REGION Network 21
   RUNG wire#powerrail
      Contact( "Carrier_21_Status.9" )
      Coil( "EMS".Carrier[21].SDC_IN.EncoderCommFault )
   END_RUNG
   // the same network as SCL:
   "EMS".Carrier[21].SDC_IN.EncoderCommFault := "Carrier_21_Status.9";
END_REGION

REGION Network 22
   RUNG wire#powerrail
      Contact( "Carrier_21_Status.10" )
      Coil( "EMS".Carrier[21].SDC_IN.DriveCommFault )
   END_RUNG
   // the same network as SCL:
   "EMS".Carrier[21].SDC_IN.DriveCommFault := "Carrier_21_Status.10";
END_REGION

REGION Network 23
   RUNG wire#powerrail
      Contact( "Carrier_21_Status.11" )
      Coil( "EMS".Carrier[21].SDC_IN.HMICommFault )
   END_RUNG
   // the same network as SCL:
   "EMS".Carrier[21].SDC_IN.HMICommFault := "Carrier_21_Status.11";
END_REGION

REGION Network 24
   RUNG wire#powerrail
      Contact( "Carrier_21_Status.2" )
      Coil( "EMS".Carrier[21].SDC_IN.AutoMode )
   END_RUNG
   RUNG wire#powerrail
      Contact( "Carrier_21_Status.1" )
      Coil( "EMS".Carrier[21].SDC_IN.ManualMode )
   END_RUNG
   // the same network as SCL:
   "EMS".Carrier[21].SDC_IN.AutoMode := "Carrier_21_Status.2";
   "EMS".Carrier[21].SDC_IN.ManualMode := "Carrier_21_Status.1";
END_REGION

REGION Network 25
   Label( C21_Comm_Fault )
   RUNG wire#powerrail
      Coil( "SectionComment" )
   END_RUNG
   // the same network as SCL:
   C21_Comm_Fault:
   "SectionComment" := TRUE;
END_REGION

REGION Network 26
   // **********************************************************************************************************************
   // 
   // Carrier 22 I-Device Data Transfer Interlocks from Carrier to SDC
   // 
   // **********************************************************************************************************************
   RUNG wire#powerrail
      Coil( "SectionComment" )
   END_RUNG
   // the same network as SCL:
   "SectionComment" := TRUE;
END_REGION

REGION Network 27
   RUNG wire#powerrail
      { S7_Templates := "SrcType := Word" } NE_Contact(in1 := "Carrier_22_CarrierNumber", in2 := 0)
      Move(in := "Carrier_22_CarrierNumber", out1 => "EMS".Carrier[22].SDC_IN.CarrierNumber)
   END_RUNG
   // the same network as SCL:
   IF "Carrier_22_CarrierNumber" <> 0 THEN
       "EMS".Carrier[22].SDC_IN.CarrierNumber := "Carrier_22_CarrierNumber";
   END_IF;
END_REGION

REGION Network 28
   RUNG wire#powerrail
      { S7_Templates := "SrcType := DWord" } NE_Contact(in1 := "Carrier_22_CarrierPosition", in2 := 0)
      Move(in := "Carrier_22_CarrierPosition", out1 => "EMS".Carrier[22].SDC_IN.CarrierPosition)
   END_RUNG
   // the same network as SCL:
   IF "Carrier_22_CarrierPosition" <> 0 THEN
       "EMS".Carrier[22].SDC_IN.CarrierPosition := "Carrier_22_CarrierPosition";
   END_IF;
END_REGION

REGION Network 29
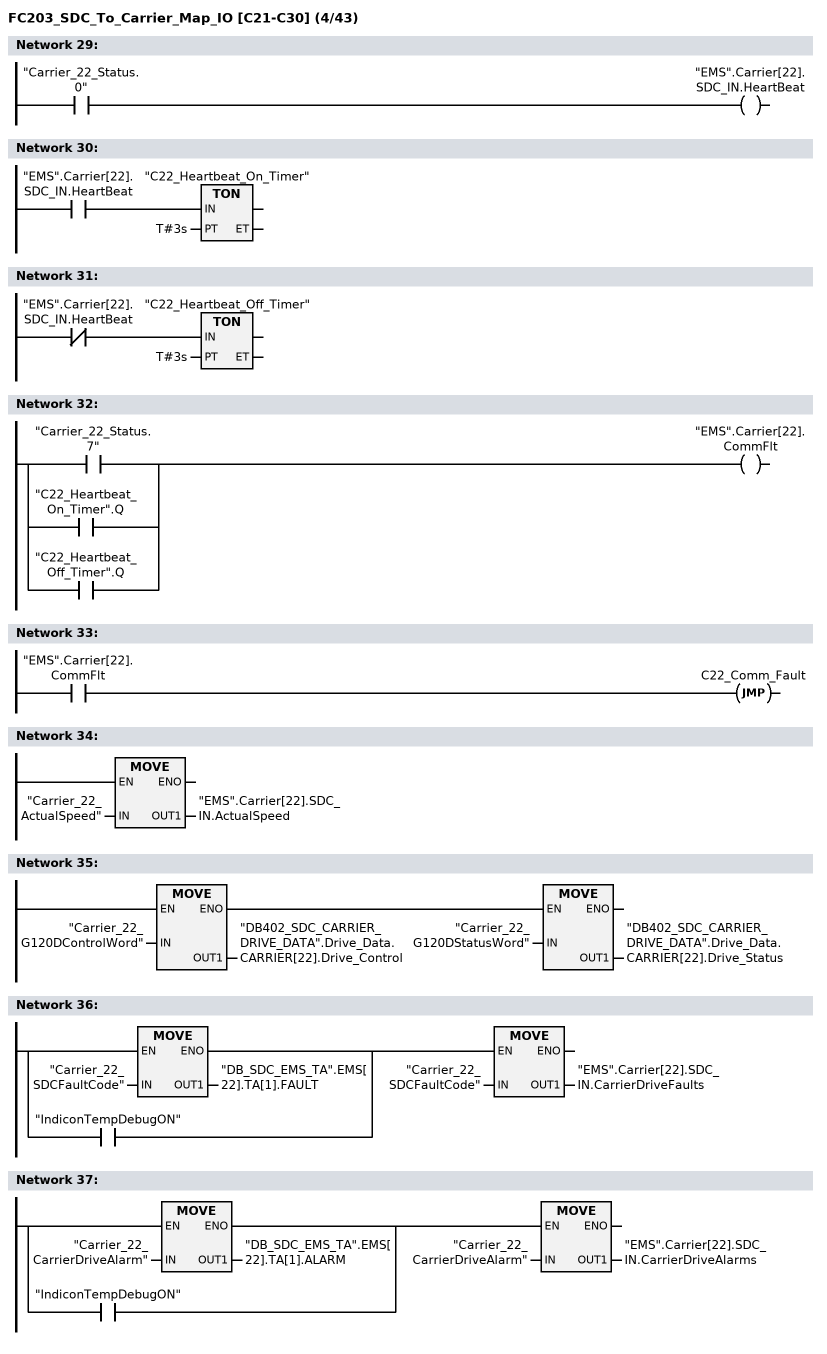
   RUNG wire#powerrail
      Contact( "Carrier_22_Status.0" )
      Coil( "EMS".Carrier[22].SDC_IN.HeartBeat )
   END_RUNG
   // the same network as SCL:
   "EMS".Carrier[22].SDC_IN.HeartBeat := "Carrier_22_Status.0";
END_REGION

REGION Network 30
   "C22_Heartbeat_On_Timer".TON(IN := "EMS".Carrier[22].SDC_IN.HeartBeat, PT := T#3s);
END_REGION

REGION Network 31
   "C22_Heartbeat_Off_Timer".TON(IN := NOT "EMS".Carrier[22].SDC_IN.HeartBeat, PT := T#3s);
END_REGION

REGION Network 32
   RUNG wire#powerrail
      Contact( "Carrier_22_Status.7" )
      wire#w1
      Coil( "EMS".Carrier[22].CommFlt )
   END_RUNG
   RUNG wire#powerrail
      Contact( "C22_Heartbeat_On_Timer".Q )
   END_RUNG wire#w1
   RUNG wire#powerrail
      Contact( "C22_Heartbeat_Off_Timer".Q )
   END_RUNG wire#w1
   // the same network as SCL:
   "EMS".Carrier[22].CommFlt := "Carrier_22_Status.7" OR "C22_Heartbeat_On_Timer".Q OR "C22_Heartbeat_Off_Timer".Q;
END_REGION

REGION Network 33
   RUNG wire#powerrail
      Contact( "EMS".Carrier[22].CommFlt )
      JumpCoil( C22_Comm_Fault )
   END_RUNG
   // the same network as SCL:
   IF "EMS".Carrier[22].CommFlt THEN GOTO C22_Comm_Fault; END_IF;
END_REGION

REGION Network 34
   RUNG wire#powerrail
      Move(in := "Carrier_22_ActualSpeed", out1 => "EMS".Carrier[22].SDC_IN.ActualSpeed)
   END_RUNG
   // the same network as SCL:
   "EMS".Carrier[22].SDC_IN.ActualSpeed := "Carrier_22_ActualSpeed";
END_REGION

REGION Network 35
   RUNG wire#powerrail
      Move(in := "Carrier_22_G120DControlWord", out1 => "DB402_SDC_CARRIER_DRIVE_DATA".Drive_Data.CARRIER[22].Drive_Control)
      Move(in := "Carrier_22_G120DStatusWord", out1 => "DB402_SDC_CARRIER_DRIVE_DATA".Drive_Data.CARRIER[22].Drive_Status)
   END_RUNG
   // the same network as SCL:
   "DB402_SDC_CARRIER_DRIVE_DATA".Drive_Data.CARRIER[22].Drive_Control := "Carrier_22_G120DControlWord";
   "DB402_SDC_CARRIER_DRIVE_DATA".Drive_Data.CARRIER[22].Drive_Status := "Carrier_22_G120DStatusWord";
END_REGION

REGION Network 36
   RUNG wire#powerrail
      Move(in := "Carrier_22_SDCFaultCode", out1 => "DB_SDC_EMS_TA".EMS[22].TA[1].FAULT)
      wire#w1
      Move(in := "Carrier_22_SDCFaultCode", out1 => "EMS".Carrier[22].SDC_IN.CarrierDriveFaults)
   END_RUNG
   RUNG wire#powerrail
      Contact( "IndiconTempDebugON" )
   END_RUNG wire#w1
   // the same network as SCL:
   "DB_SDC_EMS_TA".EMS[22].TA[1].FAULT := "Carrier_22_SDCFaultCode";
   IF TRUE OR "IndiconTempDebugON" THEN
       "EMS".Carrier[22].SDC_IN.CarrierDriveFaults := "Carrier_22_SDCFaultCode";
   END_IF;
END_REGION

REGION Network 37
   RUNG wire#powerrail
      Move(in := "Carrier_22_CarrierDriveAlarm", out1 => "DB_SDC_EMS_TA".EMS[22].TA[1].ALARM)
      wire#w1
      Move(in := "Carrier_22_CarrierDriveAlarm", out1 => "EMS".Carrier[22].SDC_IN.CarrierDriveAlarms)
   END_RUNG
   RUNG wire#powerrail
      Contact( "IndiconTempDebugON" )
   END_RUNG wire#w1
   // the same network as SCL:
   "DB_SDC_EMS_TA".EMS[22].TA[1].ALARM := "Carrier_22_CarrierDriveAlarm";
   IF TRUE OR "IndiconTempDebugON" THEN
       "EMS".Carrier[22].SDC_IN.CarrierDriveAlarms := "Carrier_22_CarrierDriveAlarm";
   END_IF;
END_REGION

REGION Network 38
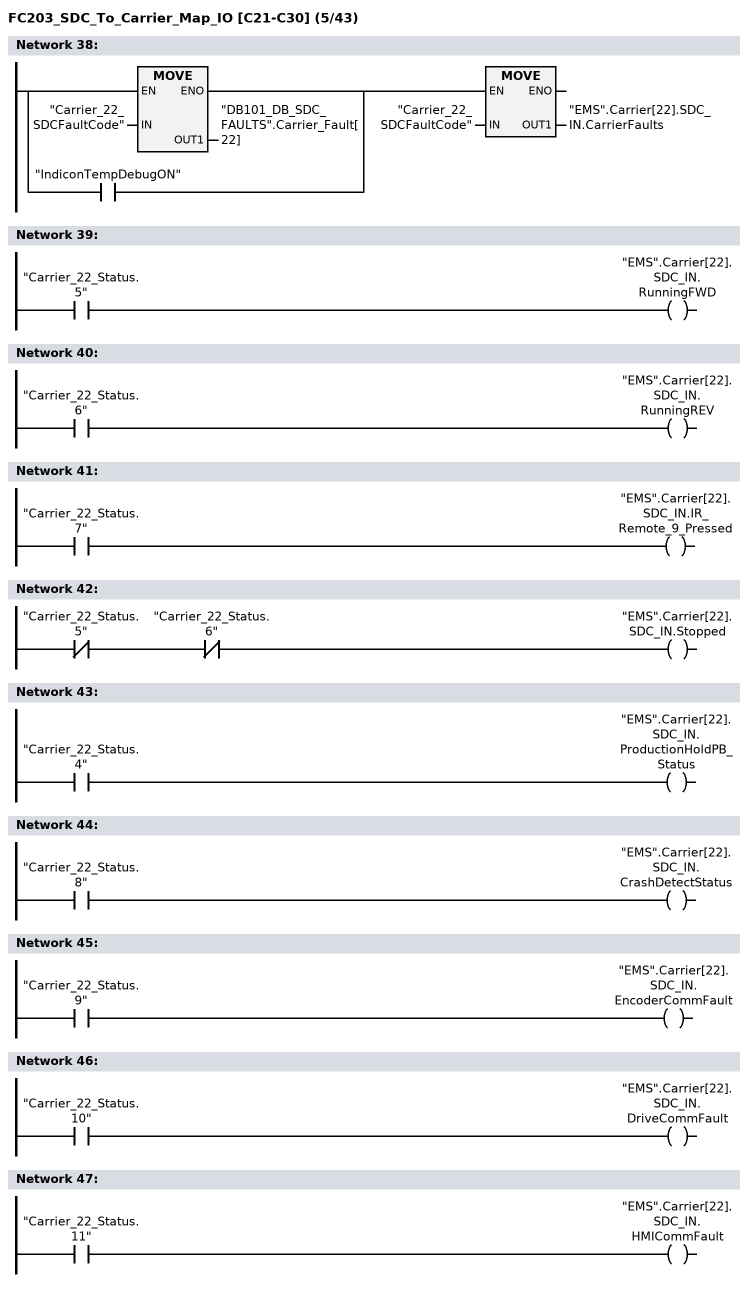
   RUNG wire#powerrail
      Move(in := "Carrier_22_SDCFaultCode", out1 => "DB101_DB_SDC_FAULTS".Carrier_Fault[22])
      wire#w1
      Move(in := "Carrier_22_SDCFaultCode", out1 => "EMS".Carrier[22].SDC_IN.CarrierFaults)
   END_RUNG
   RUNG wire#powerrail
      Contact( "IndiconTempDebugON" )
   END_RUNG wire#w1
   // the same network as SCL:
   "DB101_DB_SDC_FAULTS".Carrier_Fault[22] := "Carrier_22_SDCFaultCode";
   IF TRUE OR "IndiconTempDebugON" THEN
       "EMS".Carrier[22].SDC_IN.CarrierFaults := "Carrier_22_SDCFaultCode";
   END_IF;
END_REGION

REGION Network 39
   RUNG wire#powerrail
      Contact( "Carrier_22_Status.5" )
      Coil( "EMS".Carrier[22].SDC_IN.RunningFWD )
   END_RUNG
   // the same network as SCL:
   "EMS".Carrier[22].SDC_IN.RunningFWD := "Carrier_22_Status.5";
END_REGION

REGION Network 40
   RUNG wire#powerrail
      Contact( "Carrier_22_Status.6" )
      Coil( "EMS".Carrier[22].SDC_IN.RunningREV )
   END_RUNG
   // the same network as SCL:
   "EMS".Carrier[22].SDC_IN.RunningREV := "Carrier_22_Status.6";
END_REGION

REGION Network 41
   RUNG wire#powerrail
      Contact( "Carrier_22_Status.7" )
      Coil( "EMS".Carrier[22].SDC_IN.IR_Remote_9_Pressed )
   END_RUNG
   // the same network as SCL:
   "EMS".Carrier[22].SDC_IN.IR_Remote_9_Pressed := "Carrier_22_Status.7";
END_REGION

REGION Network 42
   RUNG wire#powerrail
      I_Contact( "Carrier_22_Status.5" )
      I_Contact( "Carrier_22_Status.6" )
      Coil( "EMS".Carrier[22].SDC_IN.Stopped )
   END_RUNG
   // the same network as SCL:
   "EMS".Carrier[22].SDC_IN.Stopped := NOT "Carrier_22_Status.5" AND NOT "Carrier_22_Status.6";
END_REGION

REGION Network 43
   RUNG wire#powerrail
      Contact( "Carrier_22_Status.4" )
      Coil( "EMS".Carrier[22].SDC_IN.ProductionHoldPB_Status )
   END_RUNG
   // the same network as SCL:
   "EMS".Carrier[22].SDC_IN.ProductionHoldPB_Status := "Carrier_22_Status.4";
END_REGION

REGION Network 44
   RUNG wire#powerrail
      Contact( "Carrier_22_Status.8" )
      Coil( "EMS".Carrier[22].SDC_IN.CrashDetectStatus )
   END_RUNG
   // the same network as SCL:
   "EMS".Carrier[22].SDC_IN.CrashDetectStatus := "Carrier_22_Status.8";
END_REGION

REGION Network 45
   RUNG wire#powerrail
      Contact( "Carrier_22_Status.9" )
      Coil( "EMS".Carrier[22].SDC_IN.EncoderCommFault )
   END_RUNG
   // the same network as SCL:
   "EMS".Carrier[22].SDC_IN.EncoderCommFault := "Carrier_22_Status.9";
END_REGION

REGION Network 46
   RUNG wire#powerrail
      Contact( "Carrier_22_Status.10" )
      Coil( "EMS".Carrier[22].SDC_IN.DriveCommFault )
   END_RUNG
   // the same network as SCL:
   "EMS".Carrier[22].SDC_IN.DriveCommFault := "Carrier_22_Status.10";
END_REGION

REGION Network 47
   RUNG wire#powerrail
      Contact( "Carrier_22_Status.11" )
      Coil( "EMS".Carrier[22].SDC_IN.HMICommFault )
   END_RUNG
   // the same network as SCL:
   "EMS".Carrier[22].SDC_IN.HMICommFault := "Carrier_22_Status.11";
END_REGION

REGION Network 48
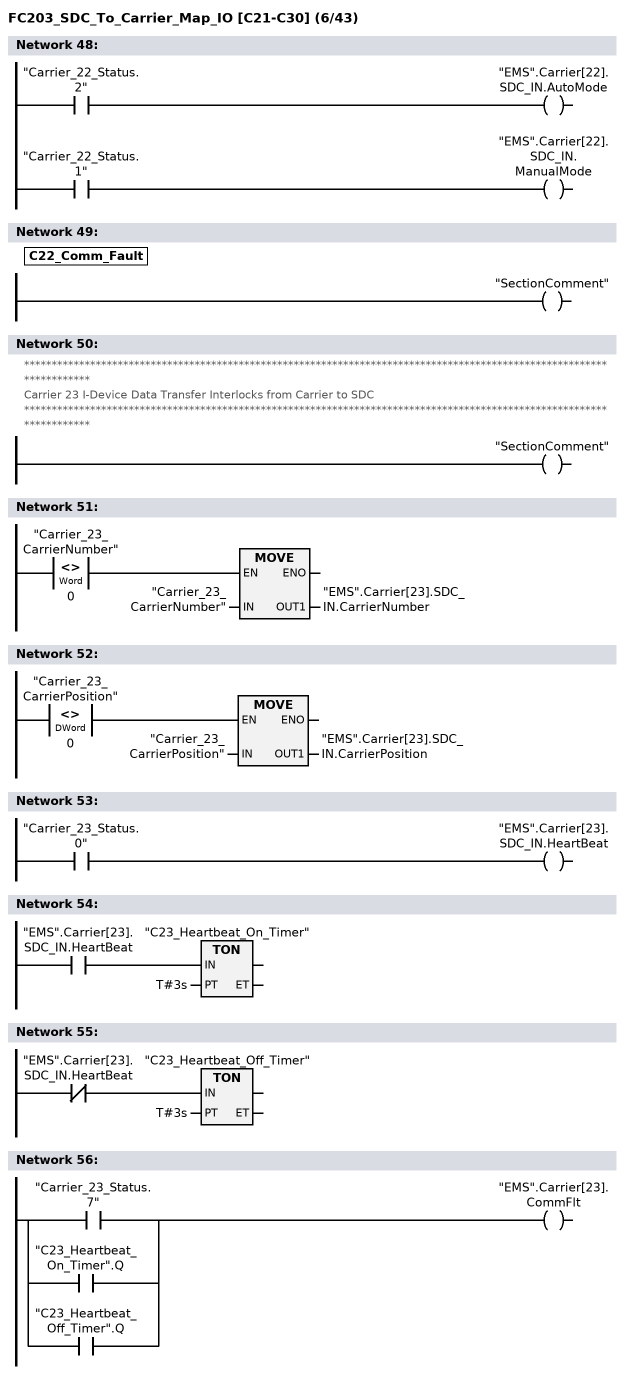
   RUNG wire#powerrail
      Contact( "Carrier_22_Status.2" )
      Coil( "EMS".Carrier[22].SDC_IN.AutoMode )
   END_RUNG
   RUNG wire#powerrail
      Contact( "Carrier_22_Status.1" )
      Coil( "EMS".Carrier[22].SDC_IN.ManualMode )
   END_RUNG
   // the same network as SCL:
   "EMS".Carrier[22].SDC_IN.AutoMode := "Carrier_22_Status.2";
   "EMS".Carrier[22].SDC_IN.ManualMode := "Carrier_22_Status.1";
END_REGION

REGION Network 49
   Label( C22_Comm_Fault )
   RUNG wire#powerrail
      Coil( "SectionComment" )
   END_RUNG
   // the same network as SCL:
   C22_Comm_Fault:
   "SectionComment" := TRUE;
END_REGION

REGION Network 50
   // **********************************************************************************************************************
   // 
   // Carrier 23 I-Device Data Transfer Interlocks from Carrier to SDC
   // 
   // **********************************************************************************************************************
   RUNG wire#powerrail
      Coil( "SectionComment" )
   END_RUNG
   // the same network as SCL:
   "SectionComment" := TRUE;
END_REGION

REGION Network 51
   RUNG wire#powerrail
      { S7_Templates := "SrcType := Word" } NE_Contact(in1 := "Carrier_23_CarrierNumber", in2 := 0)
      Move(in := "Carrier_23_CarrierNumber", out1 => "EMS".Carrier[23].SDC_IN.CarrierNumber)
   END_RUNG
   // the same network as SCL:
   IF "Carrier_23_CarrierNumber" <> 0 THEN
       "EMS".Carrier[23].SDC_IN.CarrierNumber := "Carrier_23_CarrierNumber";
   END_IF;
END_REGION

REGION Network 52
   RUNG wire#powerrail
      { S7_Templates := "SrcType := DWord" } NE_Contact(in1 := "Carrier_23_CarrierPosition", in2 := 0)
      Move(in := "Carrier_23_CarrierPosition", out1 => "EMS".Carrier[23].SDC_IN.CarrierPosition)
   END_RUNG
   // the same network as SCL:
   IF "Carrier_23_CarrierPosition" <> 0 THEN
       "EMS".Carrier[23].SDC_IN.CarrierPosition := "Carrier_23_CarrierPosition";
   END_IF;
END_REGION

REGION Network 53
   RUNG wire#powerrail
      Contact( "Carrier_23_Status.0" )
      Coil( "EMS".Carrier[23].SDC_IN.HeartBeat )
   END_RUNG
   // the same network as SCL:
   "EMS".Carrier[23].SDC_IN.HeartBeat := "Carrier_23_Status.0";
END_REGION

REGION Network 54
   "C23_Heartbeat_On_Timer".TON(IN := "EMS".Carrier[23].SDC_IN.HeartBeat, PT := T#3s);
END_REGION

REGION Network 55
   "C23_Heartbeat_Off_Timer".TON(IN := NOT "EMS".Carrier[23].SDC_IN.HeartBeat, PT := T#3s);
END_REGION

REGION Network 56
   RUNG wire#powerrail
      Contact( "Carrier_23_Status.7" )
      wire#w1
      Coil( "EMS".Carrier[23].CommFlt )
   END_RUNG
   RUNG wire#powerrail
      Contact( "C23_Heartbeat_On_Timer".Q )
   END_RUNG wire#w1
   RUNG wire#powerrail
      Contact( "C23_Heartbeat_Off_Timer".Q )
   END_RUNG wire#w1
   // the same network as SCL:
   "EMS".Carrier[23].CommFlt := "Carrier_23_Status.7" OR "C23_Heartbeat_On_Timer".Q OR "C23_Heartbeat_Off_Timer".Q;
END_REGION

REGION Network 57
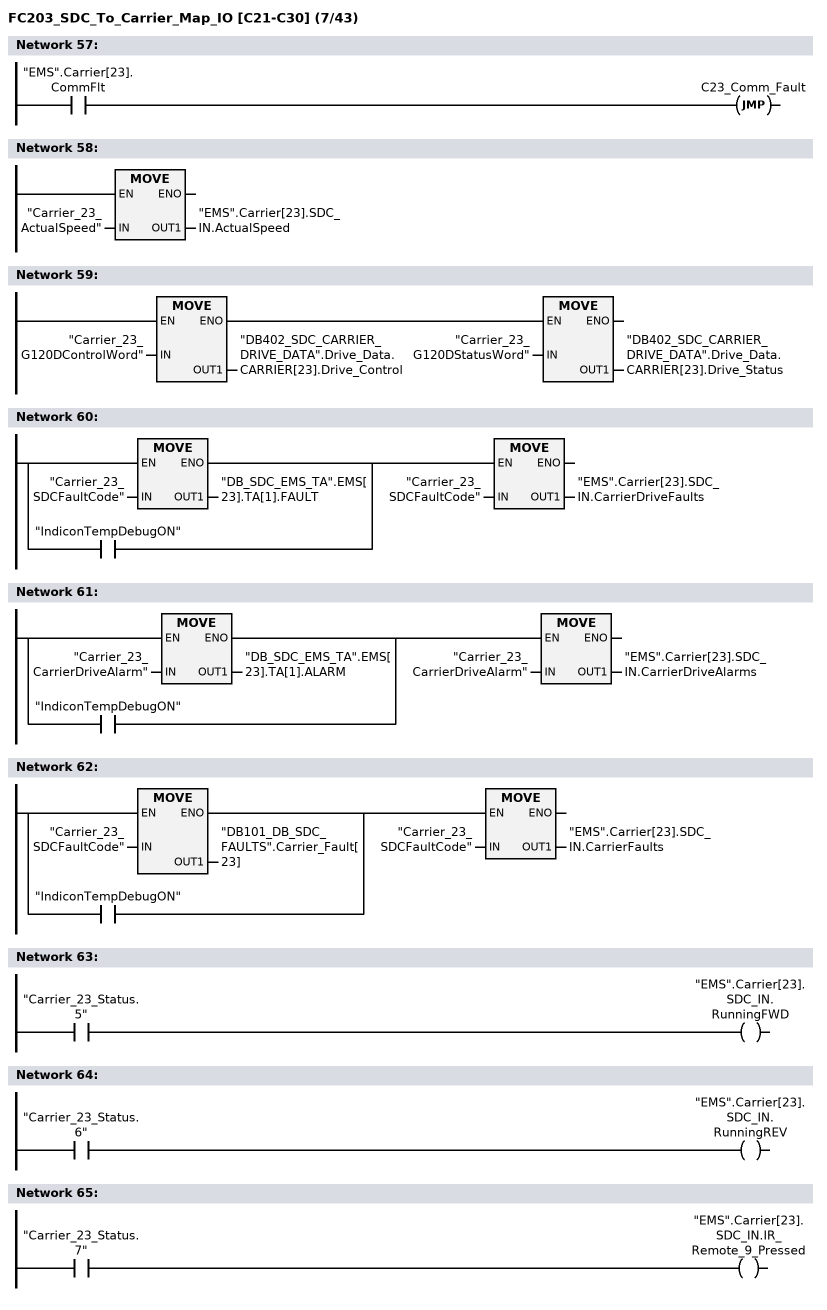
   RUNG wire#powerrail
      Contact( "EMS".Carrier[23].CommFlt )
      JumpCoil( C23_Comm_Fault )
   END_RUNG
   // the same network as SCL:
   IF "EMS".Carrier[23].CommFlt THEN GOTO C23_Comm_Fault; END_IF;
END_REGION

REGION Network 58
   RUNG wire#powerrail
      Move(in := "Carrier_23_ActualSpeed", out1 => "EMS".Carrier[23].SDC_IN.ActualSpeed)
   END_RUNG
   // the same network as SCL:
   "EMS".Carrier[23].SDC_IN.ActualSpeed := "Carrier_23_ActualSpeed";
END_REGION

REGION Network 59
   RUNG wire#powerrail
      Move(in := "Carrier_23_G120DControlWord", out1 => "DB402_SDC_CARRIER_DRIVE_DATA".Drive_Data.CARRIER[23].Drive_Control)
      Move(in := "Carrier_23_G120DStatusWord", out1 => "DB402_SDC_CARRIER_DRIVE_DATA".Drive_Data.CARRIER[23].Drive_Status)
   END_RUNG
   // the same network as SCL:
   "DB402_SDC_CARRIER_DRIVE_DATA".Drive_Data.CARRIER[23].Drive_Control := "Carrier_23_G120DControlWord";
   "DB402_SDC_CARRIER_DRIVE_DATA".Drive_Data.CARRIER[23].Drive_Status := "Carrier_23_G120DStatusWord";
END_REGION

REGION Network 60
   RUNG wire#powerrail
      Move(in := "Carrier_23_SDCFaultCode", out1 => "DB_SDC_EMS_TA".EMS[23].TA[1].FAULT)
      wire#w1
      Move(in := "Carrier_23_SDCFaultCode", out1 => "EMS".Carrier[23].SDC_IN.CarrierDriveFaults)
   END_RUNG
   RUNG wire#powerrail
      Contact( "IndiconTempDebugON" )
   END_RUNG wire#w1
   // the same network as SCL:
   "DB_SDC_EMS_TA".EMS[23].TA[1].FAULT := "Carrier_23_SDCFaultCode";
   IF TRUE OR "IndiconTempDebugON" THEN
       "EMS".Carrier[23].SDC_IN.CarrierDriveFaults := "Carrier_23_SDCFaultCode";
   END_IF;
END_REGION

REGION Network 61
   RUNG wire#powerrail
      Move(in := "Carrier_23_CarrierDriveAlarm", out1 => "DB_SDC_EMS_TA".EMS[23].TA[1].ALARM)
      wire#w1
      Move(in := "Carrier_23_CarrierDriveAlarm", out1 => "EMS".Carrier[23].SDC_IN.CarrierDriveAlarms)
   END_RUNG
   RUNG wire#powerrail
      Contact( "IndiconTempDebugON" )
   END_RUNG wire#w1
   // the same network as SCL:
   "DB_SDC_EMS_TA".EMS[23].TA[1].ALARM := "Carrier_23_CarrierDriveAlarm";
   IF TRUE OR "IndiconTempDebugON" THEN
       "EMS".Carrier[23].SDC_IN.CarrierDriveAlarms := "Carrier_23_CarrierDriveAlarm";
   END_IF;
END_REGION

REGION Network 62
   RUNG wire#powerrail
      Move(in := "Carrier_23_SDCFaultCode", out1 => "DB101_DB_SDC_FAULTS".Carrier_Fault[23])
      wire#w1
      Move(in := "Carrier_23_SDCFaultCode", out1 => "EMS".Carrier[23].SDC_IN.CarrierFaults)
   END_RUNG
   RUNG wire#powerrail
      Contact( "IndiconTempDebugON" )
   END_RUNG wire#w1
   // the same network as SCL:
   "DB101_DB_SDC_FAULTS".Carrier_Fault[23] := "Carrier_23_SDCFaultCode";
   IF TRUE OR "IndiconTempDebugON" THEN
       "EMS".Carrier[23].SDC_IN.CarrierFaults := "Carrier_23_SDCFaultCode";
   END_IF;
END_REGION

REGION Network 63
   RUNG wire#powerrail
      Contact( "Carrier_23_Status.5" )
      Coil( "EMS".Carrier[23].SDC_IN.RunningFWD )
   END_RUNG
   // the same network as SCL:
   "EMS".Carrier[23].SDC_IN.RunningFWD := "Carrier_23_Status.5";
END_REGION

REGION Network 64
   RUNG wire#powerrail
      Contact( "Carrier_23_Status.6" )
      Coil( "EMS".Carrier[23].SDC_IN.RunningREV )
   END_RUNG
   // the same network as SCL:
   "EMS".Carrier[23].SDC_IN.RunningREV := "Carrier_23_Status.6";
END_REGION

REGION Network 65
   RUNG wire#powerrail
      Contact( "Carrier_23_Status.7" )
      Coil( "EMS".Carrier[23].SDC_IN.IR_Remote_9_Pressed )
   END_RUNG
   // the same network as SCL:
   "EMS".Carrier[23].SDC_IN.IR_Remote_9_Pressed := "Carrier_23_Status.7";
END_REGION

REGION Network 66
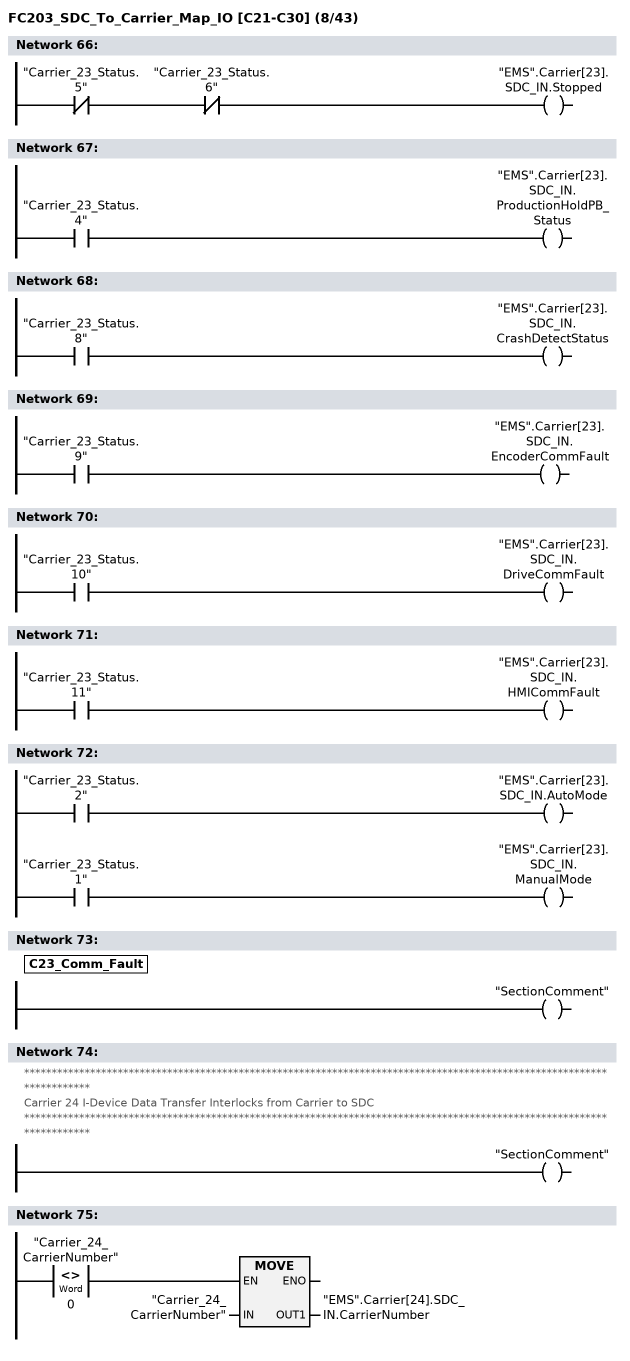
   RUNG wire#powerrail
      I_Contact( "Carrier_23_Status.5" )
      I_Contact( "Carrier_23_Status.6" )
      Coil( "EMS".Carrier[23].SDC_IN.Stopped )
   END_RUNG
   // the same network as SCL:
   "EMS".Carrier[23].SDC_IN.Stopped := NOT "Carrier_23_Status.5" AND NOT "Carrier_23_Status.6";
END_REGION

REGION Network 67
   RUNG wire#powerrail
      Contact( "Carrier_23_Status.4" )
      Coil( "EMS".Carrier[23].SDC_IN.ProductionHoldPB_Status )
   END_RUNG
   // the same network as SCL:
   "EMS".Carrier[23].SDC_IN.ProductionHoldPB_Status := "Carrier_23_Status.4";
END_REGION

REGION Network 68
   RUNG wire#powerrail
      Contact( "Carrier_23_Status.8" )
      Coil( "EMS".Carrier[23].SDC_IN.CrashDetectStatus )
   END_RUNG
   // the same network as SCL:
   "EMS".Carrier[23].SDC_IN.CrashDetectStatus := "Carrier_23_Status.8";
END_REGION

REGION Network 69
   RUNG wire#powerrail
      Contact( "Carrier_23_Status.9" )
      Coil( "EMS".Carrier[23].SDC_IN.EncoderCommFault )
   END_RUNG
   // the same network as SCL:
   "EMS".Carrier[23].SDC_IN.EncoderCommFault := "Carrier_23_Status.9";
END_REGION

REGION Network 70
   RUNG wire#powerrail
      Contact( "Carrier_23_Status.10" )
      Coil( "EMS".Carrier[23].SDC_IN.DriveCommFault )
   END_RUNG
   // the same network as SCL:
   "EMS".Carrier[23].SDC_IN.DriveCommFault := "Carrier_23_Status.10";
END_REGION

REGION Network 71
   RUNG wire#powerrail
      Contact( "Carrier_23_Status.11" )
      Coil( "EMS".Carrier[23].SDC_IN.HMICommFault )
   END_RUNG
   // the same network as SCL:
   "EMS".Carrier[23].SDC_IN.HMICommFault := "Carrier_23_Status.11";
END_REGION

REGION Network 72
   RUNG wire#powerrail
      Contact( "Carrier_23_Status.2" )
      Coil( "EMS".Carrier[23].SDC_IN.AutoMode )
   END_RUNG
   RUNG wire#powerrail
      Contact( "Carrier_23_Status.1" )
      Coil( "EMS".Carrier[23].SDC_IN.ManualMode )
   END_RUNG
   // the same network as SCL:
   "EMS".Carrier[23].SDC_IN.AutoMode := "Carrier_23_Status.2";
   "EMS".Carrier[23].SDC_IN.ManualMode := "Carrier_23_Status.1";
END_REGION

REGION Network 73
   Label( C23_Comm_Fault )
   RUNG wire#powerrail
      Coil( "SectionComment" )
   END_RUNG
   // the same network as SCL:
   C23_Comm_Fault:
   "SectionComment" := TRUE;
END_REGION

REGION Network 74
   // **********************************************************************************************************************
   // 
   // Carrier 24 I-Device Data Transfer Interlocks from Carrier to SDC
   // 
   // **********************************************************************************************************************
   RUNG wire#powerrail
      Coil( "SectionComment" )
   END_RUNG
   // the same network as SCL:
   "SectionComment" := TRUE;
END_REGION

REGION Network 75
   RUNG wire#powerrail
      { S7_Templates := "SrcType := Word" } NE_Contact(in1 := "Carrier_24_CarrierNumber", in2 := 0)
      Move(in := "Carrier_24_CarrierNumber", out1 => "EMS".Carrier[24].SDC_IN.CarrierNumber)
   END_RUNG
   // the same network as SCL:
   IF "Carrier_24_CarrierNumber" <> 0 THEN
       "EMS".Carrier[24].SDC_IN.CarrierNumber := "Carrier_24_CarrierNumber";
   END_IF;
END_REGION

REGION Network 76
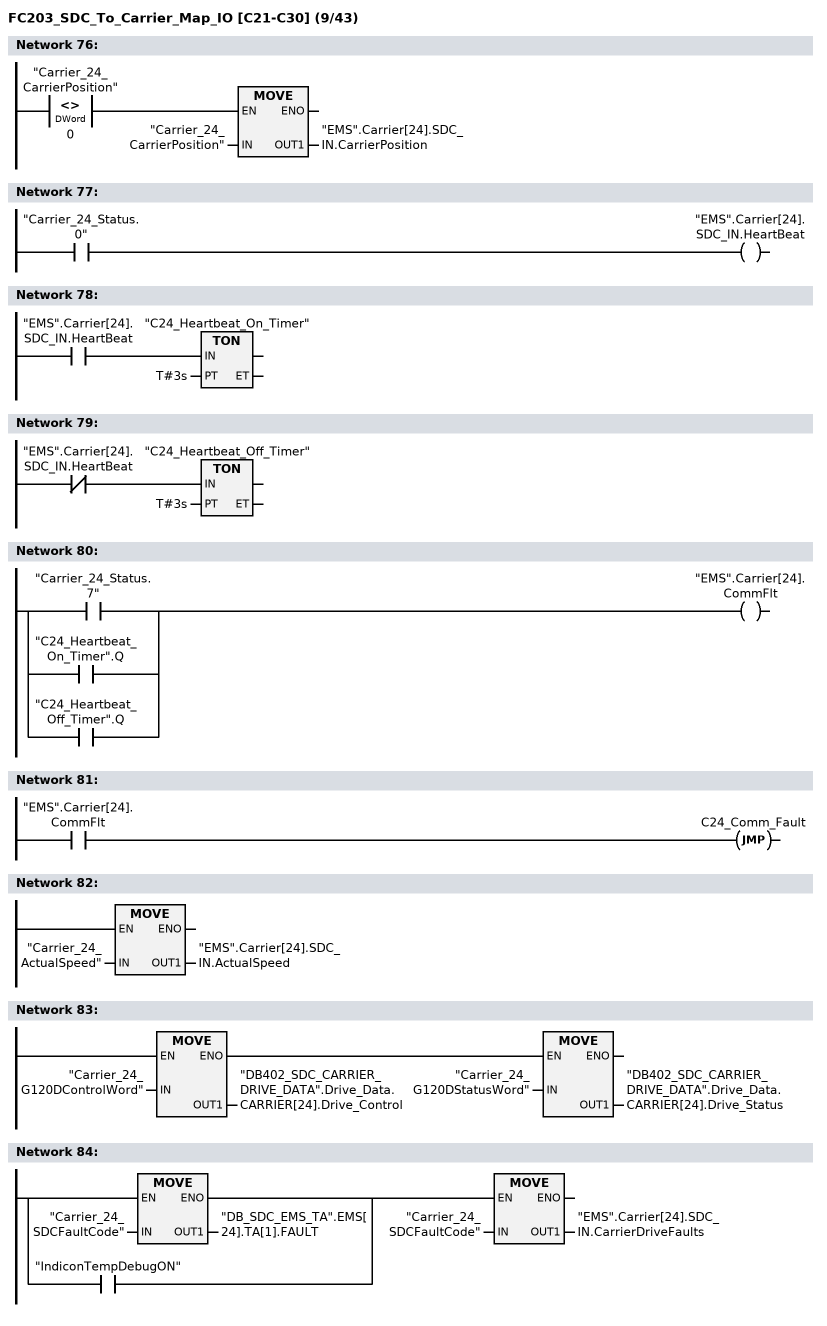
   RUNG wire#powerrail
      { S7_Templates := "SrcType := DWord" } NE_Contact(in1 := "Carrier_24_CarrierPosition", in2 := 0)
      Move(in := "Carrier_24_CarrierPosition", out1 => "EMS".Carrier[24].SDC_IN.CarrierPosition)
   END_RUNG
   // the same network as SCL:
   IF "Carrier_24_CarrierPosition" <> 0 THEN
       "EMS".Carrier[24].SDC_IN.CarrierPosition := "Carrier_24_CarrierPosition";
   END_IF;
END_REGION

REGION Network 77
   RUNG wire#powerrail
      Contact( "Carrier_24_Status.0" )
      Coil( "EMS".Carrier[24].SDC_IN.HeartBeat )
   END_RUNG
   // the same network as SCL:
   "EMS".Carrier[24].SDC_IN.HeartBeat := "Carrier_24_Status.0";
END_REGION

REGION Network 78
   "C24_Heartbeat_On_Timer".TON(IN := "EMS".Carrier[24].SDC_IN.HeartBeat, PT := T#3s);
END_REGION

REGION Network 79
   "C24_Heartbeat_Off_Timer".TON(IN := NOT "EMS".Carrier[24].SDC_IN.HeartBeat, PT := T#3s);
END_REGION

REGION Network 80
   RUNG wire#powerrail
      Contact( "Carrier_24_Status.7" )
      wire#w1
      Coil( "EMS".Carrier[24].CommFlt )
   END_RUNG
   RUNG wire#powerrail
      Contact( "C24_Heartbeat_On_Timer".Q )
   END_RUNG wire#w1
   RUNG wire#powerrail
      Contact( "C24_Heartbeat_Off_Timer".Q )
   END_RUNG wire#w1
   // the same network as SCL:
   "EMS".Carrier[24].CommFlt := "Carrier_24_Status.7" OR "C24_Heartbeat_On_Timer".Q OR "C24_Heartbeat_Off_Timer".Q;
END_REGION

REGION Network 81
   RUNG wire#powerrail
      Contact( "EMS".Carrier[24].CommFlt )
      JumpCoil( C24_Comm_Fault )
   END_RUNG
   // the same network as SCL:
   IF "EMS".Carrier[24].CommFlt THEN GOTO C24_Comm_Fault; END_IF;
END_REGION

REGION Network 82
   RUNG wire#powerrail
      Move(in := "Carrier_24_ActualSpeed", out1 => "EMS".Carrier[24].SDC_IN.ActualSpeed)
   END_RUNG
   // the same network as SCL:
   "EMS".Carrier[24].SDC_IN.ActualSpeed := "Carrier_24_ActualSpeed";
END_REGION

REGION Network 83
   RUNG wire#powerrail
      Move(in := "Carrier_24_G120DControlWord", out1 => "DB402_SDC_CARRIER_DRIVE_DATA".Drive_Data.CARRIER[24].Drive_Control)
      Move(in := "Carrier_24_G120DStatusWord", out1 => "DB402_SDC_CARRIER_DRIVE_DATA".Drive_Data.CARRIER[24].Drive_Status)
   END_RUNG
   // the same network as SCL:
   "DB402_SDC_CARRIER_DRIVE_DATA".Drive_Data.CARRIER[24].Drive_Control := "Carrier_24_G120DControlWord";
   "DB402_SDC_CARRIER_DRIVE_DATA".Drive_Data.CARRIER[24].Drive_Status := "Carrier_24_G120DStatusWord";
END_REGION

REGION Network 84
   RUNG wire#powerrail
      Move(in := "Carrier_24_SDCFaultCode", out1 => "DB_SDC_EMS_TA".EMS[24].TA[1].FAULT)
      wire#w1
      Move(in := "Carrier_24_SDCFaultCode", out1 => "EMS".Carrier[24].SDC_IN.CarrierDriveFaults)
   END_RUNG
   RUNG wire#powerrail
      Contact( "IndiconTempDebugON" )
   END_RUNG wire#w1
   // the same network as SCL:
   "DB_SDC_EMS_TA".EMS[24].TA[1].FAULT := "Carrier_24_SDCFaultCode";
   IF TRUE OR "IndiconTempDebugON" THEN
       "EMS".Carrier[24].SDC_IN.CarrierDriveFaults := "Carrier_24_SDCFaultCode";
   END_IF;
END_REGION

REGION Network 85
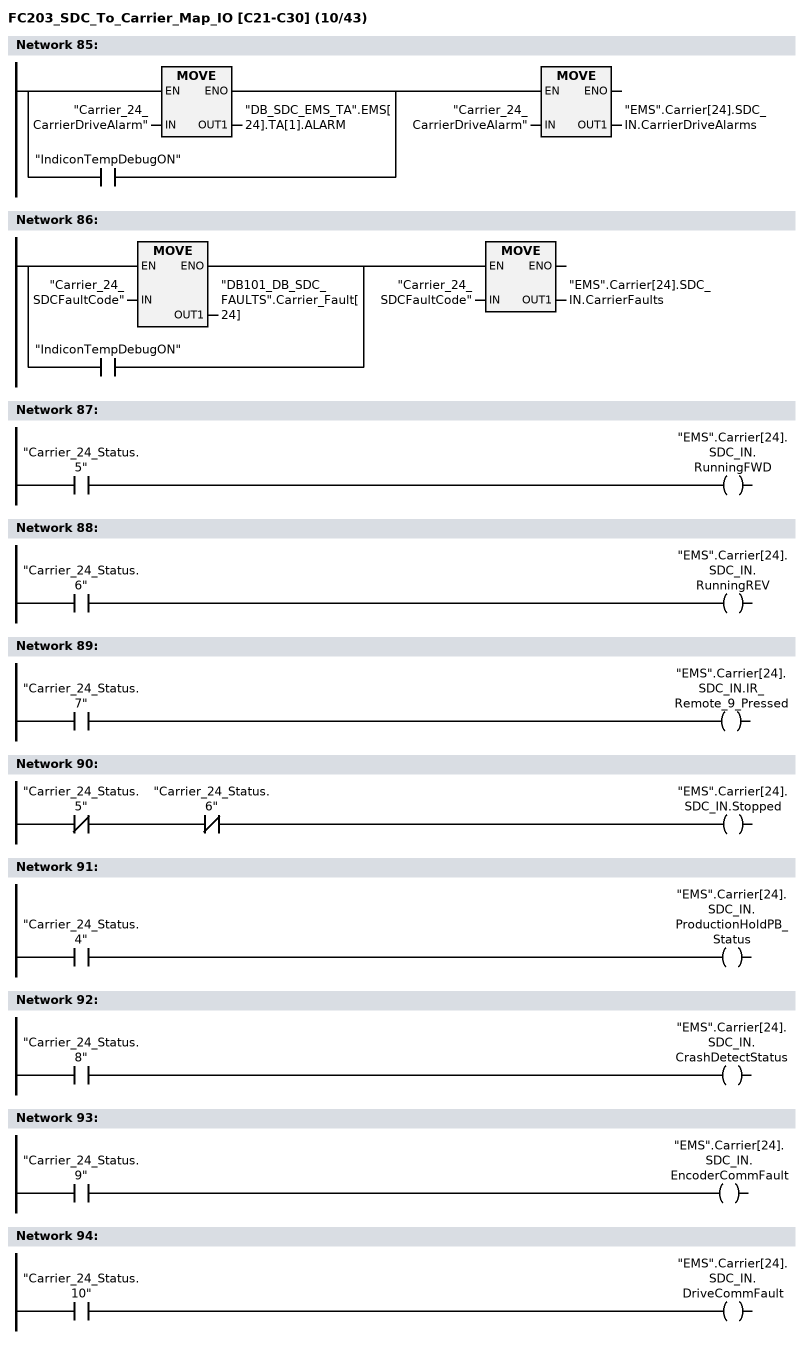
   RUNG wire#powerrail
      Move(in := "Carrier_24_CarrierDriveAlarm", out1 => "DB_SDC_EMS_TA".EMS[24].TA[1].ALARM)
      wire#w1
      Move(in := "Carrier_24_CarrierDriveAlarm", out1 => "EMS".Carrier[24].SDC_IN.CarrierDriveAlarms)
   END_RUNG
   RUNG wire#powerrail
      Contact( "IndiconTempDebugON" )
   END_RUNG wire#w1
   // the same network as SCL:
   "DB_SDC_EMS_TA".EMS[24].TA[1].ALARM := "Carrier_24_CarrierDriveAlarm";
   IF TRUE OR "IndiconTempDebugON" THEN
       "EMS".Carrier[24].SDC_IN.CarrierDriveAlarms := "Carrier_24_CarrierDriveAlarm";
   END_IF;
END_REGION

REGION Network 86
   RUNG wire#powerrail
      Move(in := "Carrier_24_SDCFaultCode", out1 => "DB101_DB_SDC_FAULTS".Carrier_Fault[24])
      wire#w1
      Move(in := "Carrier_24_SDCFaultCode", out1 => "EMS".Carrier[24].SDC_IN.CarrierFaults)
   END_RUNG
   RUNG wire#powerrail
      Contact( "IndiconTempDebugON" )
   END_RUNG wire#w1
   // the same network as SCL:
   "DB101_DB_SDC_FAULTS".Carrier_Fault[24] := "Carrier_24_SDCFaultCode";
   IF TRUE OR "IndiconTempDebugON" THEN
       "EMS".Carrier[24].SDC_IN.CarrierFaults := "Carrier_24_SDCFaultCode";
   END_IF;
END_REGION

REGION Network 87
   RUNG wire#powerrail
      Contact( "Carrier_24_Status.5" )
      Coil( "EMS".Carrier[24].SDC_IN.RunningFWD )
   END_RUNG
   // the same network as SCL:
   "EMS".Carrier[24].SDC_IN.RunningFWD := "Carrier_24_Status.5";
END_REGION

REGION Network 88
   RUNG wire#powerrail
      Contact( "Carrier_24_Status.6" )
      Coil( "EMS".Carrier[24].SDC_IN.RunningREV )
   END_RUNG
   // the same network as SCL:
   "EMS".Carrier[24].SDC_IN.RunningREV := "Carrier_24_Status.6";
END_REGION

REGION Network 89
   RUNG wire#powerrail
      Contact( "Carrier_24_Status.7" )
      Coil( "EMS".Carrier[24].SDC_IN.IR_Remote_9_Pressed )
   END_RUNG
   // the same network as SCL:
   "EMS".Carrier[24].SDC_IN.IR_Remote_9_Pressed := "Carrier_24_Status.7";
END_REGION

REGION Network 90
   RUNG wire#powerrail
      I_Contact( "Carrier_24_Status.5" )
      I_Contact( "Carrier_24_Status.6" )
      Coil( "EMS".Carrier[24].SDC_IN.Stopped )
   END_RUNG
   // the same network as SCL:
   "EMS".Carrier[24].SDC_IN.Stopped := NOT "Carrier_24_Status.5" AND NOT "Carrier_24_Status.6";
END_REGION

REGION Network 91
   RUNG wire#powerrail
      Contact( "Carrier_24_Status.4" )
      Coil( "EMS".Carrier[24].SDC_IN.ProductionHoldPB_Status )
   END_RUNG
   // the same network as SCL:
   "EMS".Carrier[24].SDC_IN.ProductionHoldPB_Status := "Carrier_24_Status.4";
END_REGION

REGION Network 92
   RUNG wire#powerrail
      Contact( "Carrier_24_Status.8" )
      Coil( "EMS".Carrier[24].SDC_IN.CrashDetectStatus )
   END_RUNG
   // the same network as SCL:
   "EMS".Carrier[24].SDC_IN.CrashDetectStatus := "Carrier_24_Status.8";
END_REGION

REGION Network 93
   RUNG wire#powerrail
      Contact( "Carrier_24_Status.9" )
      Coil( "EMS".Carrier[24].SDC_IN.EncoderCommFault )
   END_RUNG
   // the same network as SCL:
   "EMS".Carrier[24].SDC_IN.EncoderCommFault := "Carrier_24_Status.9";
END_REGION

REGION Network 94
   RUNG wire#powerrail
      Contact( "Carrier_24_Status.10" )
      Coil( "EMS".Carrier[24].SDC_IN.DriveCommFault )
   END_RUNG
   // the same network as SCL:
   "EMS".Carrier[24].SDC_IN.DriveCommFault := "Carrier_24_Status.10";
END_REGION

REGION Network 95
